   IF #COM_RST              // полный сброс
   THEN
       #LMNR_SIM:=#LMNRSVAL;
       #QLMNUP:=0;
       #QLMNDN:=0;
       #PV:=0.0;
       #ER:=0.0;
       #LMNRS_ON:=0;
       #LMNRSVAL:=0.0;
       #LMNR_SIM:=0.0;
       #sFbPVal:=0.0;
       #sThrOn:=0.0;
       #siImpAus:=0;
       #stImpDauer:=T#0MS;
       #stPausDauer:=T#0MS;
   ELSE
       #Istwert:=INT_TO_REAL(WORD_TO_INT(#PV_PER))*3.616898e-003;
       #Istwert:=#Istwert*#PV_FAC+#PV_OFF;
       IF NOT #PVPER_ON THEN #Istwert:=#PV_IN; END_IF;
       #PV:=#Istwert;
       #ErKp:=#SP_INT-#PV;
       IF    #ErKp < (-#DEADB_W) THEN  #ER:=#ErKp+#DEADB_W;
       ELSIF #ErKp>#DEADB_W      THEN  #ER:=#ErKp-#DEADB_W;
       ELSE  #ER:=0.0; END_IF;
       #ErKp:=#ER*#GAIN;
       #rCycle:=DINT_TO_REAL(TIME_TO_DINT(#CYCLE))/1000.0;
       #rTi:=DINT_TO_REAL(TIME_TO_DINT(#TI))/1000.0;
       IF #rTi<#rCycle*0.5 THEN #rTi:=#rCycle*0.5; END_IF;
       #rMtrTm:=DINT_TO_REAL(TIME_TO_DINT(#MTR_TM))/1000.0;
       #Hvar:=#rTi-ABS(0.01*#ErKp*#rMtrTm);
       IF #Hvar<(#rTi*0.1)THEN #rTi:=#rTi*0.1; ELSE #rTi:=#Hvar; END_IF; 
       IF #LMNS_ON
       THEN
           #sFbPVal:=0.0;
       ELSE 
           IF #siImpAus<>0
           THEN 
               #dInteg:=DINT_TO_REAL(INT_TO_DINT(#siImpAus))*#rCycle/#rMtrTm;
           ELSE
               IF (#ErKp>0.0 AND #LMNR_HS) OR (#ErKp<0.0 AND #LMNR_LS) OR (#TI=T#0MS) 
               THEN
                   #dInteg:=0.0;
               ELSE   
                   #dInteg := (-#ErKp)*#rCycle/#rTi;
               END_IF;
           END_IF;
           #sFbPVal:=#sFbPVal+#dInteg;
           IF #TI=T#0MS
           THEN 
               IF    #sFbPVal>100.0 THEN #sFbPVal:=100.0;
               ELSIF #sFbPVal<0.0   THEN #sFbPVal:=0.0;
               END_IF;
           END_IF;   
       END_IF;       
       #dThrStIn:=#ErKp-#sFbPVal+#DISV;
       #AdapIn1:=#ErKp;
       #AdapIn2:=#sFbPVal;
       #rThrOff:=55.0/#rMtrTm*#rCycle;
       IF #PULSE_TM>#CYCLE
       THEN 
       #Hvar:=DINT_TO_REAL(TIME_TO_DINT(#PULSE_TM))/1000.0;
       ELSE
       #Hvar:=#rCycle;
       END_IF;
       #Hvar:=100.0*#Hvar/#rMtrTm;
       IF NOT(#LMNR_HS OR #LMNR_LS)
       THEN
           IF NOT (#QLMNUP OR #QLMNDN)
           THEN
               IF #TI<>T#0MS
               THEN
                   IF ABS(#AdapIn1)<ABS(#AdapIn2)
                   THEN
                       #sThrOn:=#AdapIn1;
                   ELSE    
                       #sThrOn:=#AdapIn2;
                   END_IF;
               ELSE
                   IF #Istwert=0.0
                   THEN
                       #sThrOn:=#Hvar;
                   ELSE
                       #sThrOn:=ABS(#ErKp)*0.5;
                   END_IF;
               END_IF;
               IF #sThrOn>10.0 THEN #sThrOn:=10.0; END_IF;
               IF #sThrOn<#Hvar THEN #sThrOn:=#Hvar; END_IF;            
           END_IF;           
       ELSE 
           #sThrOn:=#Hvar;
       END_IF;     
       IF (#siImpAus=100 AND #dThrStIn>#rThrOff) OR (#dThrStIn>=#sThrOn)             THEN #iImpEin:=100;
       ELSIF (#siImpAus=-100 AND #dThrStIn<(-#rThrOff)) OR (#dThrStIn<=(-#sThrOn))   THEN #iImpEin:=-100;
       ELSE                                                                          #iImpEin:=0;     
       END_IF;
       IF  #LMNS_ON
       THEN
           IF #LMNUP XOR #LMNDN 
           THEN
               IF #LMNUP
               THEN
                   #iImpEin:=100;
               ELSE
                   #iImpEin:=-100;
               END_IF;
           ELSE
               #iImpEin:=0;
           END_IF;
       END_IF;   
       IF (#iImpEin=100 AND #LMNR_HS) OR (#iImpEin=-100 AND #LMNR_LS) THEN #iImpEin:=0; END_IF;
       IF (#siImpAus=-100 AND #iImpEin=100) OR (#siImpAus=100 AND #iImpEin=-100)THEN #iImpEin:=0; END_IF;
       IF #siImpAus<>#iImpEin
       THEN
           IF #iImpEin=0
           THEN
               IF #stImpDauer<=T#0MS
               THEN
                   #siImpAus:=0;
                   #stPausDauer:=#BREAK_TM;
               END_IF;
           ELSE
               #siImpAus:=#iImpEin;
               #stImpDauer:=#PULSE_TM;
           END_IF;
       END_IF;
       IF #stImpDauer>T#0MS
       THEN
       #stImpDauer:=#stImpDauer-#CYCLE;
       ELSE
       #stImpDauer:=T#0MS;
       END_IF;
       IF #stPausDauer>T#0MS
       THEN
       #stPausDauer:=#stPausDauer-#CYCLE;
       ELSE 
       #stPausDauer:=T#0MS;
       END_IF;
       IF ((#siImpAus=100) AND #LMNR_HS) OR ((#siImpAus=-100) AND #LMNR_LS)
       THEN
         #siImpAus:=0;
         #stImpDauer:=T#0MS;
       END_IF;
       IF NOT #LMNRS_ON
       THEN
           #LmnrSim:=#LMNRSVAL;
       ELSE
           #LmnrSim:=DINT_TO_REAL(INT_TO_DINT(#siImpAus))*#rCycle/#rMtrTm+#LMNR_SIM;
           IF #LmnrSim>=100.0
           THEN
               #LmnrSim:=100.0;
           ELSIF  #LmnrSim<=0.0
           THEN
               #LmnrSim:=0.0;
           END_IF;
       END_IF;
       #LMNR_SIM:=#LmnrSim;
       IF #siImpAus=0
       THEN
              #QLMNUP:=0;
              #QLMNDN:=0;
       ELSIF #siImpAus=100
       THEN
           #QLMNUP:=1;
                 #QLMNDN:=0;
       ELSE
              #QLMNUP:=0;
              #QLMNDN:=1;
       END_IF;
   END_IF;
END_FUNCTION_BLOCK

FUNCTION "03_FC_PID" : Void   // FC3, LAD
{ S7_Optimized_Access := 'FALSE' }
VERSION : 0.1
BEGIN

REGION Network 1
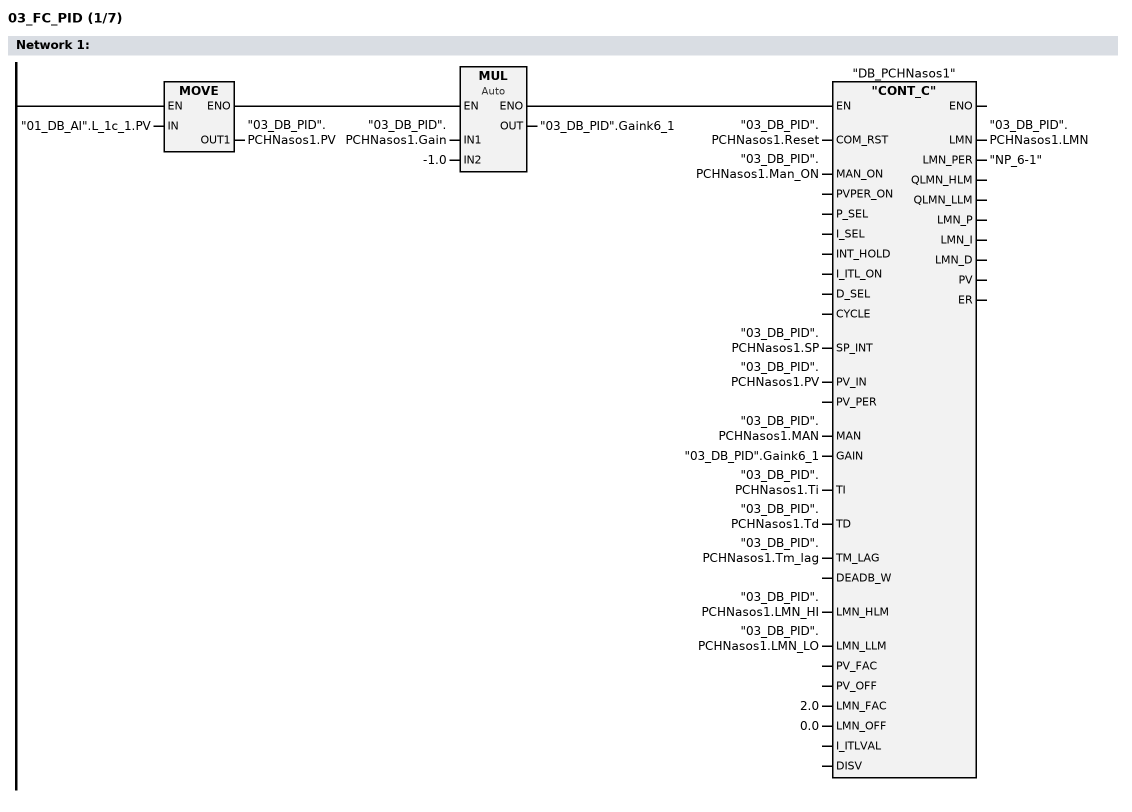
   RUNG wire#powerrail
      Move(in := "01_DB_AI".L_1c_1.PV, out1 => "03_DB_PID".PCHNasos1.PV)
      Mul(in1 := "03_DB_PID".PCHNasos1.Gain, in2 := -1.0, out => "03_DB_PID".Gaink6_1)
      "DB_PCHNasos1"(COM_RST := "03_DB_PID".PCHNasos1.Reset, MAN_ON := "03_DB_PID".PCHNasos1.Man_ON, PVPER_ON :=, P_SEL :=, I_SEL :=, INT_HOLD :=, I_ITL_ON :=, D_SEL :=, CYCLE :=, SP_INT := "03_DB_PID".PCHNasos1.SP, PV_IN := "03_DB_PID".PCHNasos1.PV, PV_PER :=, MAN := "03_DB_PID".PCHNasos1.MAN, GAIN := "03_DB_PID".Gaink6_1, TI := "03_DB_PID".PCHNasos1.Ti, TD := "03_DB_PID".PCHNasos1.Td, TM_LAG := "03_DB_PID".PCHNasos1.Tm_lag, DEADB_W :=, LMN_HLM := "03_DB_PID".PCHNasos1.LMN_HI, LMN_LLM := "03_DB_PID".PCHNasos1.LMN_LO, PV_FAC :=, PV_OFF :=, LMN_FAC := 2.0, LMN_OFF := 0.0, I_ITLVAL :=, DISV :=, LMN => "03_DB_PID".PCHNasos1.LMN, LMN_PER => "NP_6-1", QLMN_HLM =>, QLMN_LLM =>, LMN_P =>, LMN_I =>, LMN_D =>, PV =>, ER =>)
   END_RUNG
   // the same network as SCL:
   "03_DB_PID".PCHNasos1.PV := "01_DB_AI".L_1c_1.PV;
   "03_DB_PID".Gaink6_1 := "03_DB_PID".PCHNasos1.Gain * (-1.0);
   "DB_PCHNasos1"(COM_RST := "03_DB_PID".PCHNasos1.Reset,   // "CONT_C"
                  MAN_ON := "03_DB_PID".PCHNasos1.Man_ON,
                  SP_INT := "03_DB_PID".PCHNasos1.SP,
                  PV_IN := "03_DB_PID".PCHNasos1.PV,
                  MAN := "03_DB_PID".PCHNasos1.MAN,
                  GAIN := "03_DB_PID".Gaink6_1,
                  TI := "03_DB_PID".PCHNasos1.Ti,
                  TD := "03_DB_PID".PCHNasos1.Td,
                  TM_LAG := "03_DB_PID".PCHNasos1.Tm_lag,
                  LMN_HLM := "03_DB_PID".PCHNasos1.LMN_HI,
                  LMN_LLM := "03_DB_PID".PCHNasos1.LMN_LO,
                  LMN_FAC := 2.0,
                  LMN_OFF := 0.0,
                  LMN => "03_DB_PID".PCHNasos1.LMN,
                  LMN_PER => "NP_6-1");
END_REGION

REGION Network 2
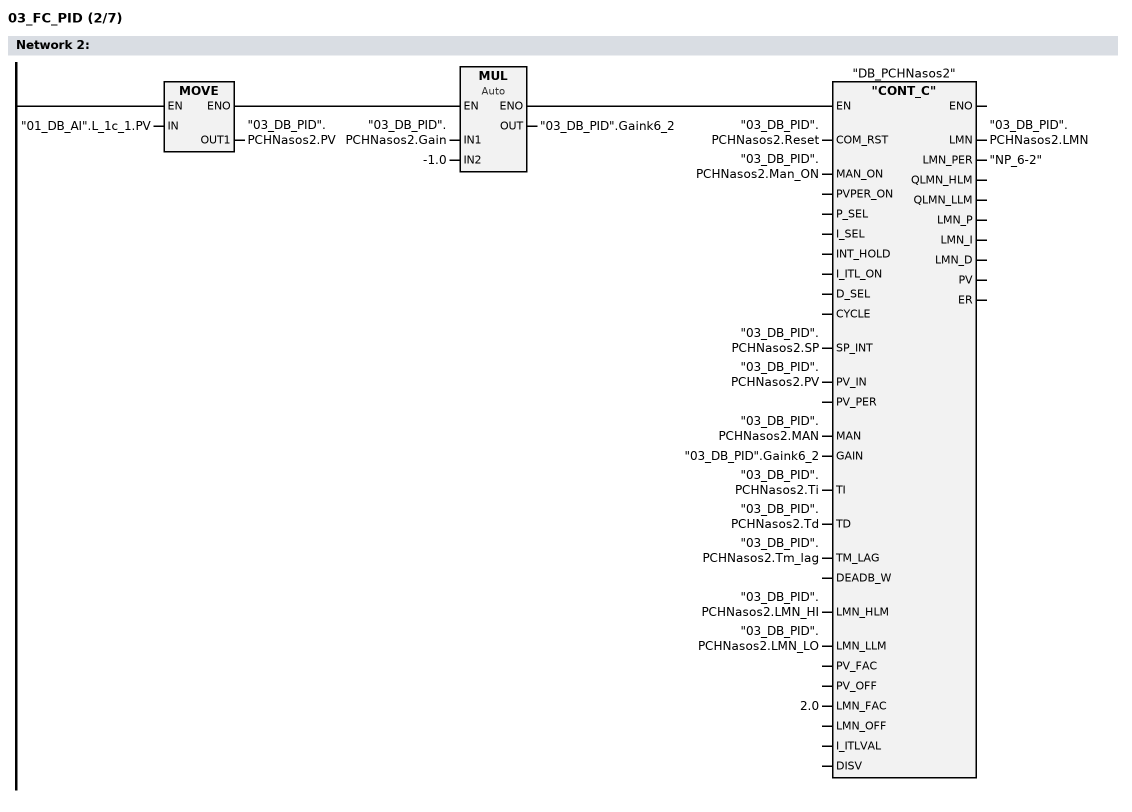
   RUNG wire#powerrail
      Move(in := "01_DB_AI".L_1c_1.PV, out1 => "03_DB_PID".PCHNasos2.PV)
      Mul(in1 := "03_DB_PID".PCHNasos2.Gain, in2 := -1.0, out => "03_DB_PID".Gaink6_2)
      "DB_PCHNasos2"(COM_RST := "03_DB_PID".PCHNasos2.Reset, MAN_ON := "03_DB_PID".PCHNasos2.Man_ON, PVPER_ON :=, P_SEL :=, I_SEL :=, INT_HOLD :=, I_ITL_ON :=, D_SEL :=, CYCLE :=, SP_INT := "03_DB_PID".PCHNasos2.SP, PV_IN := "03_DB_PID".PCHNasos2.PV, PV_PER :=, MAN := "03_DB_PID".PCHNasos2.MAN, GAIN := "03_DB_PID".Gaink6_2, TI := "03_DB_PID".PCHNasos2.Ti, TD := "03_DB_PID".PCHNasos2.Td, TM_LAG := "03_DB_PID".PCHNasos2.Tm_lag, DEADB_W :=, LMN_HLM := "03_DB_PID".PCHNasos2.LMN_HI, LMN_LLM := "03_DB_PID".PCHNasos2.LMN_LO, PV_FAC :=, PV_OFF :=, LMN_FAC := 2.0, LMN_OFF :=, I_ITLVAL :=, DISV :=, LMN => "03_DB_PID".PCHNasos2.LMN, LMN_PER => "NP_6-2", QLMN_HLM =>, QLMN_LLM =>, LMN_P =>, LMN_I =>, LMN_D =>, PV =>, ER =>)
   END_RUNG
   // the same network as SCL:
   "03_DB_PID".PCHNasos2.PV := "01_DB_AI".L_1c_1.PV;
   "03_DB_PID".Gaink6_2 := "03_DB_PID".PCHNasos2.Gain * (-1.0);
   "DB_PCHNasos2"(COM_RST := "03_DB_PID".PCHNasos2.Reset,   // "CONT_C"
                  MAN_ON := "03_DB_PID".PCHNasos2.Man_ON,
                  SP_INT := "03_DB_PID".PCHNasos2.SP,
                  PV_IN := "03_DB_PID".PCHNasos2.PV,
                  MAN := "03_DB_PID".PCHNasos2.MAN,
                  GAIN := "03_DB_PID".Gaink6_2,
                  TI := "03_DB_PID".PCHNasos2.Ti,
                  TD := "03_DB_PID".PCHNasos2.Td,
                  TM_LAG := "03_DB_PID".PCHNasos2.Tm_lag,
                  LMN_HLM := "03_DB_PID".PCHNasos2.LMN_HI,
                  LMN_LLM := "03_DB_PID".PCHNasos2.LMN_LO,
                  LMN_FAC := 2.0,
                  LMN => "03_DB_PID".PCHNasos2.LMN,
                  LMN_PER => "NP_6-2");
END_REGION

REGION Network 3
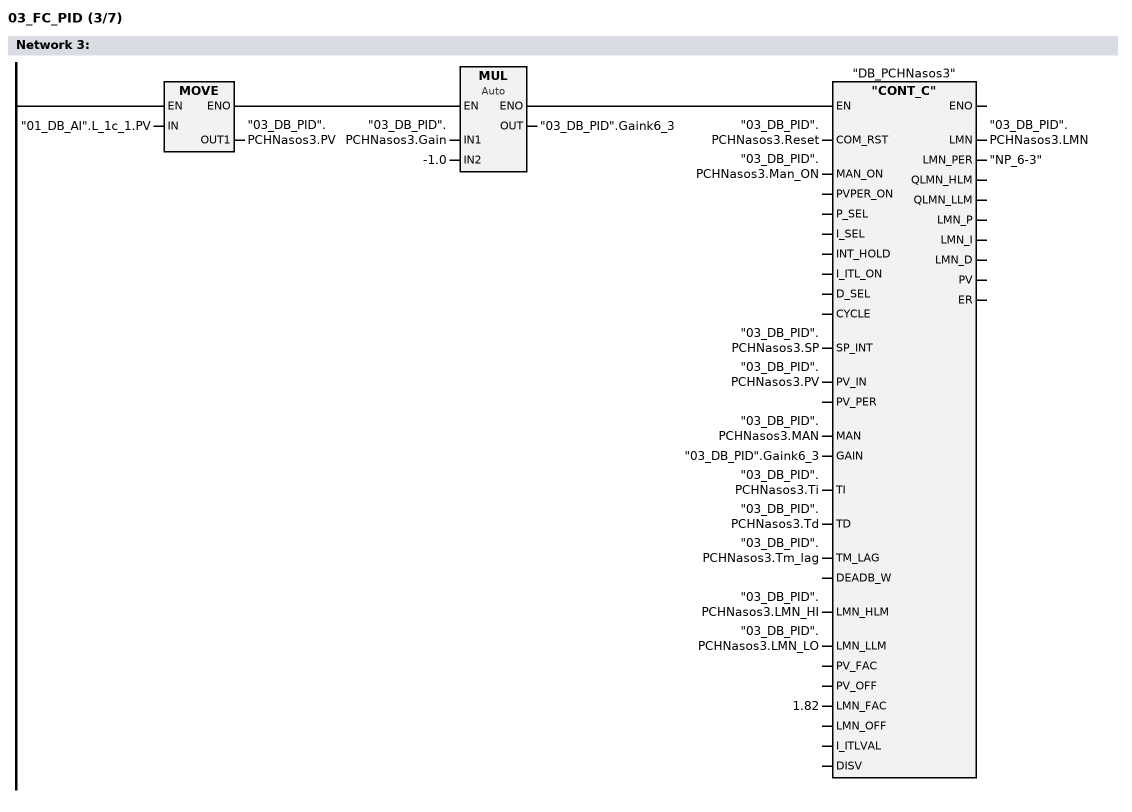
   RUNG wire#powerrail
      Move(in := "01_DB_AI".L_1c_1.PV, out1 => "03_DB_PID".PCHNasos3.PV)
      Mul(in1 := "03_DB_PID".PCHNasos3.Gain, in2 := -1.0, out => "03_DB_PID".Gaink6_3)
      "DB_PCHNasos3"(COM_RST := "03_DB_PID".PCHNasos3.Reset, MAN_ON := "03_DB_PID".PCHNasos3.Man_ON, PVPER_ON :=, P_SEL :=, I_SEL :=, INT_HOLD :=, I_ITL_ON :=, D_SEL :=, CYCLE :=, SP_INT := "03_DB_PID".PCHNasos3.SP, PV_IN := "03_DB_PID".PCHNasos3.PV, PV_PER :=, MAN := "03_DB_PID".PCHNasos3.MAN, GAIN := "03_DB_PID".Gaink6_3, TI := "03_DB_PID".PCHNasos3.Ti, TD := "03_DB_PID".PCHNasos3.Td, TM_LAG := "03_DB_PID".PCHNasos3.Tm_lag, DEADB_W :=, LMN_HLM := "03_DB_PID".PCHNasos3.LMN_HI, LMN_LLM := "03_DB_PID".PCHNasos3.LMN_LO, PV_FAC :=, PV_OFF :=, LMN_FAC := 1.82, LMN_OFF :=, I_ITLVAL :=, DISV :=, LMN => "03_DB_PID".PCHNasos3.LMN, LMN_PER => "NP_6-3", QLMN_HLM =>, QLMN_LLM =>, LMN_P =>, LMN_I =>, LMN_D =>, PV =>, ER =>)
   END_RUNG
   // the same network as SCL:
   "03_DB_PID".PCHNasos3.PV := "01_DB_AI".L_1c_1.PV;
   "03_DB_PID".Gaink6_3 := "03_DB_PID".PCHNasos3.Gain * (-1.0);
   "DB_PCHNasos3"(COM_RST := "03_DB_PID".PCHNasos3.Reset,   // "CONT_C"
                  MAN_ON := "03_DB_PID".PCHNasos3.Man_ON,
                  SP_INT := "03_DB_PID".PCHNasos3.SP,
                  PV_IN := "03_DB_PID".PCHNasos3.PV,
                  MAN := "03_DB_PID".PCHNasos3.MAN,
                  GAIN := "03_DB_PID".Gaink6_3,
                  TI := "03_DB_PID".PCHNasos3.Ti,
                  TD := "03_DB_PID".PCHNasos3.Td,
                  TM_LAG := "03_DB_PID".PCHNasos3.Tm_lag,
                  LMN_HLM := "03_DB_PID".PCHNasos3.LMN_HI,
                  LMN_LLM := "03_DB_PID".PCHNasos3.LMN_LO,
                  LMN_FAC := 1.82,
                  LMN => "03_DB_PID".PCHNasos3.LMN,
                  LMN_PER => "NP_6-3");
END_REGION

REGION Network 4
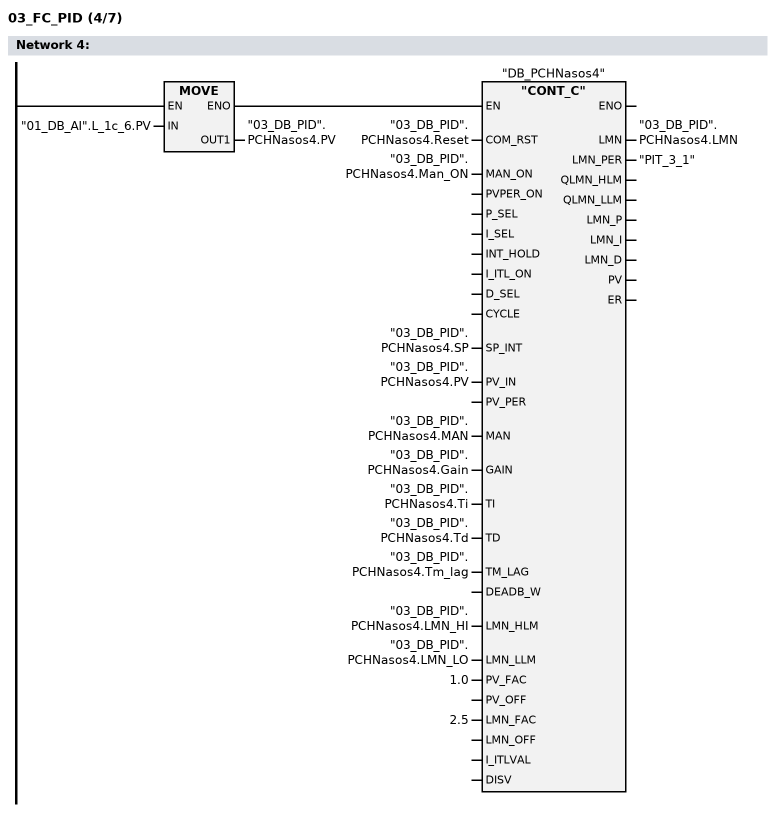
   RUNG wire#powerrail
      Move(in := "01_DB_AI".L_1c_6.PV, out1 => "03_DB_PID".PCHNasos4.PV)
      "DB_PCHNasos4"(COM_RST := "03_DB_PID".PCHNasos4.Reset, MAN_ON := "03_DB_PID".PCHNasos4.Man_ON, PVPER_ON :=, P_SEL :=, I_SEL :=, INT_HOLD :=, I_ITL_ON :=, D_SEL :=, CYCLE :=, SP_INT := "03_DB_PID".PCHNasos4.SP, PV_IN := "03_DB_PID".PCHNasos4.PV, PV_PER :=, MAN := "03_DB_PID".PCHNasos4.MAN, GAIN := "03_DB_PID".PCHNasos4.Gain, TI := "03_DB_PID".PCHNasos4.Ti, TD := "03_DB_PID".PCHNasos4.Td, TM_LAG := "03_DB_PID".PCHNasos4.Tm_lag, DEADB_W :=, LMN_HLM := "03_DB_PID".PCHNasos4.LMN_HI, LMN_LLM := "03_DB_PID".PCHNasos4.LMN_LO, PV_FAC := 1.0, PV_OFF :=, LMN_FAC := 2.5, LMN_OFF :=, I_ITLVAL :=, DISV :=, LMN => "03_DB_PID".PCHNasos4.LMN, LMN_PER => "PIT_3_1", QLMN_HLM =>, QLMN_LLM =>, LMN_P =>, LMN_I =>, LMN_D =>, PV =>, ER =>)
   END_RUNG
   // the same network as SCL:
   "03_DB_PID".PCHNasos4.PV := "01_DB_AI".L_1c_6.PV;
   "DB_PCHNasos4"(COM_RST := "03_DB_PID".PCHNasos4.Reset,   // "CONT_C"
                  MAN_ON := "03_DB_PID".PCHNasos4.Man_ON,
                  SP_INT := "03_DB_PID".PCHNasos4.SP,
                  PV_IN := "03_DB_PID".PCHNasos4.PV,
                  MAN := "03_DB_PID".PCHNasos4.MAN,
                  GAIN := "03_DB_PID".PCHNasos4.Gain,
                  TI := "03_DB_PID".PCHNasos4.Ti,
                  TD := "03_DB_PID".PCHNasos4.Td,
                  TM_LAG := "03_DB_PID".PCHNasos4.Tm_lag,
                  LMN_HLM := "03_DB_PID".PCHNasos4.LMN_HI,
                  LMN_LLM := "03_DB_PID".PCHNasos4.LMN_LO,
                  PV_FAC := 1.0,
                  LMN_FAC := 2.5,
                  LMN => "03_DB_PID".PCHNasos4.LMN,
                  LMN_PER => "PIT_3_1");
END_REGION

REGION Network 5
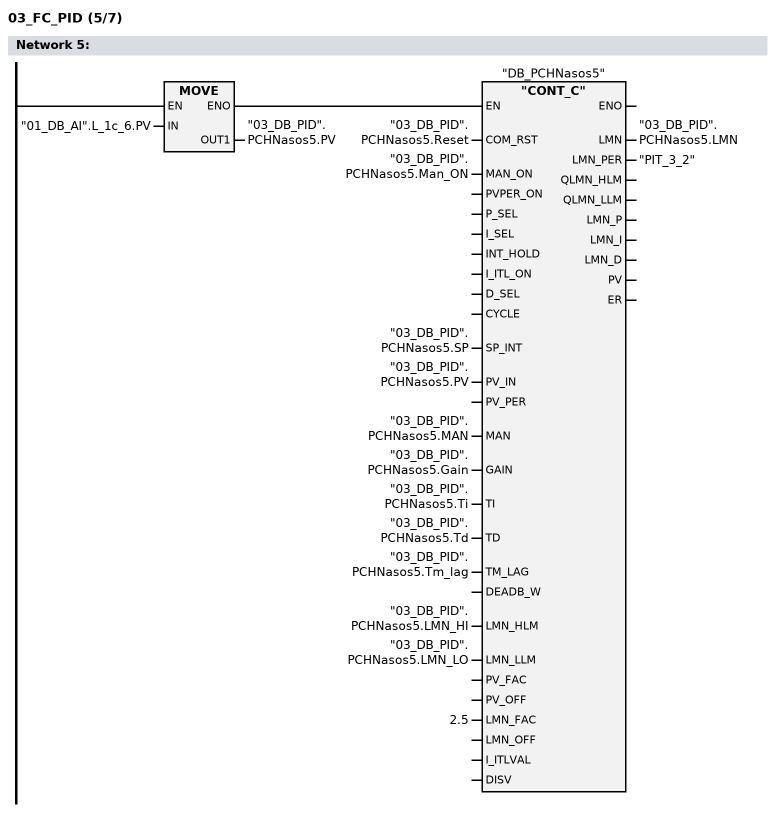
   RUNG wire#powerrail
      Move(in := "01_DB_AI".L_1c_6.PV, out1 => "03_DB_PID".PCHNasos5.PV)
      "DB_PCHNasos5"(COM_RST := "03_DB_PID".PCHNasos5.Reset, MAN_ON := "03_DB_PID".PCHNasos5.Man_ON, PVPER_ON :=, P_SEL :=, I_SEL :=, INT_HOLD :=, I_ITL_ON :=, D_SEL :=, CYCLE :=, SP_INT := "03_DB_PID".PCHNasos5.SP, PV_IN := "03_DB_PID".PCHNasos5.PV, PV_PER :=, MAN := "03_DB_PID".PCHNasos5.MAN, GAIN := "03_DB_PID".PCHNasos5.Gain, TI := "03_DB_PID".PCHNasos5.Ti, TD := "03_DB_PID".PCHNasos5.Td, TM_LAG := "03_DB_PID".PCHNasos5.Tm_lag, DEADB_W :=, LMN_HLM := "03_DB_PID".PCHNasos5.LMN_HI, LMN_LLM := "03_DB_PID".PCHNasos5.LMN_LO, PV_FAC :=, PV_OFF :=, LMN_FAC := 2.5, LMN_OFF :=, I_ITLVAL :=, DISV :=, LMN => "03_DB_PID".PCHNasos5.LMN, LMN_PER => "PIT_3_2", QLMN_HLM =>, QLMN_LLM =>, LMN_P =>, LMN_I =>, LMN_D =>, PV =>, ER =>)
   END_RUNG
   // the same network as SCL:
   "03_DB_PID".PCHNasos5.PV := "01_DB_AI".L_1c_6.PV;
   "DB_PCHNasos5"(COM_RST := "03_DB_PID".PCHNasos5.Reset,   // "CONT_C"
                  MAN_ON := "03_DB_PID".PCHNasos5.Man_ON,
                  SP_INT := "03_DB_PID".PCHNasos5.SP,
                  PV_IN := "03_DB_PID".PCHNasos5.PV,
                  MAN := "03_DB_PID".PCHNasos5.MAN,
                  GAIN := "03_DB_PID".PCHNasos5.Gain,
                  TI := "03_DB_PID".PCHNasos5.Ti,
                  TD := "03_DB_PID".PCHNasos5.Td,
                  TM_LAG := "03_DB_PID".PCHNasos5.Tm_lag,
                  LMN_HLM := "03_DB_PID".PCHNasos5.LMN_HI,
                  LMN_LLM := "03_DB_PID".PCHNasos5.LMN_LO,
                  LMN_FAC := 2.5,
                  LMN => "03_DB_PID".PCHNasos5.LMN,
                  LMN_PER => "PIT_3_2");
END_REGION

REGION Network 6
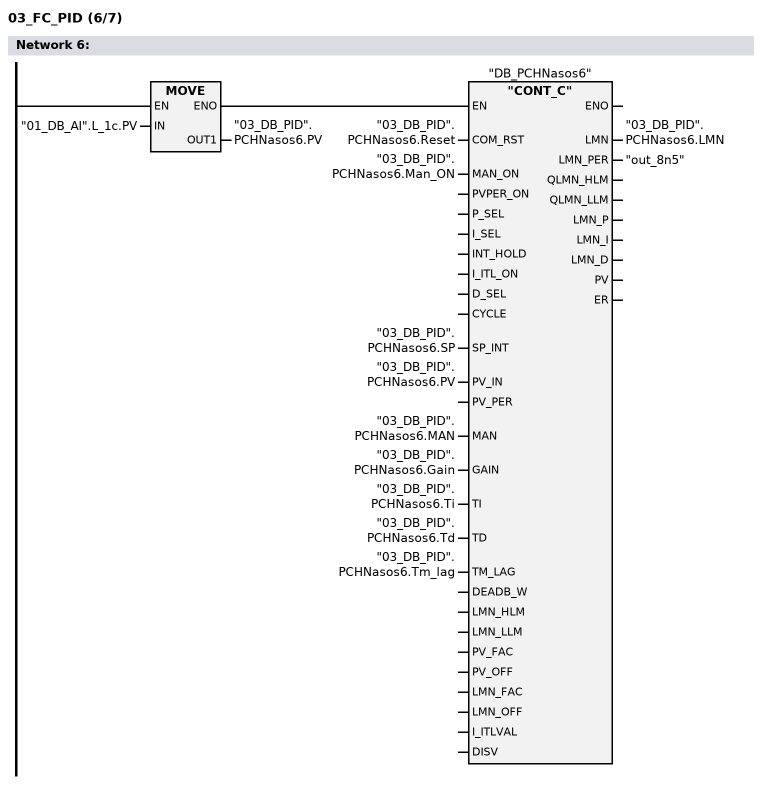
   RUNG wire#powerrail
      Move(in := "01_DB_AI".L_1c.PV, out1 => "03_DB_PID".PCHNasos6.PV)
      "DB_PCHNasos6"(COM_RST := "03_DB_PID".PCHNasos6.Reset, MAN_ON := "03_DB_PID".PCHNasos6.Man_ON, PVPER_ON :=, P_SEL :=, I_SEL :=, INT_HOLD :=, I_ITL_ON :=, D_SEL :=, CYCLE :=, SP_INT := "03_DB_PID".PCHNasos6.SP, PV_IN := "03_DB_PID".PCHNasos6.PV, PV_PER :=, MAN := "03_DB_PID".PCHNasos6.MAN, GAIN := "03_DB_PID".PCHNasos6.Gain, TI := "03_DB_PID".PCHNasos6.Ti, TD := "03_DB_PID".PCHNasos6.Td, TM_LAG := "03_DB_PID".PCHNasos6.Tm_lag, DEADB_W :=, LMN_HLM :=, LMN_LLM :=, PV_FAC :=, PV_OFF :=, LMN_FAC :=, LMN_OFF :=, I_ITLVAL :=, DISV :=, LMN => "03_DB_PID".PCHNasos6.LMN, LMN_PER => "out_8n5", QLMN_HLM =>, QLMN_LLM =>, LMN_P =>, LMN_I =>, LMN_D =>, PV =>, ER =>)
   END_RUNG
   // the same network as SCL:
   "03_DB_PID".PCHNasos6.PV := "01_DB_AI".L_1c.PV;
   "DB_PCHNasos6"(COM_RST := "03_DB_PID".PCHNasos6.Reset,   // "CONT_C"
                  MAN_ON := "03_DB_PID".PCHNasos6.Man_ON,
                  SP_INT := "03_DB_PID".PCHNasos6.SP,
                  PV_IN := "03_DB_PID".PCHNasos6.PV,
                  MAN := "03_DB_PID".PCHNasos6.MAN,
                  GAIN := "03_DB_PID".PCHNasos6.Gain,
                  TI := "03_DB_PID".PCHNasos6.Ti,
                  TD := "03_DB_PID".PCHNasos6.Td,
                  TM_LAG := "03_DB_PID".PCHNasos6.Tm_lag,
                  LMN => "03_DB_PID".PCHNasos6.LMN,
                  LMN_PER => "out_8n5");
END_REGION

REGION Network 7
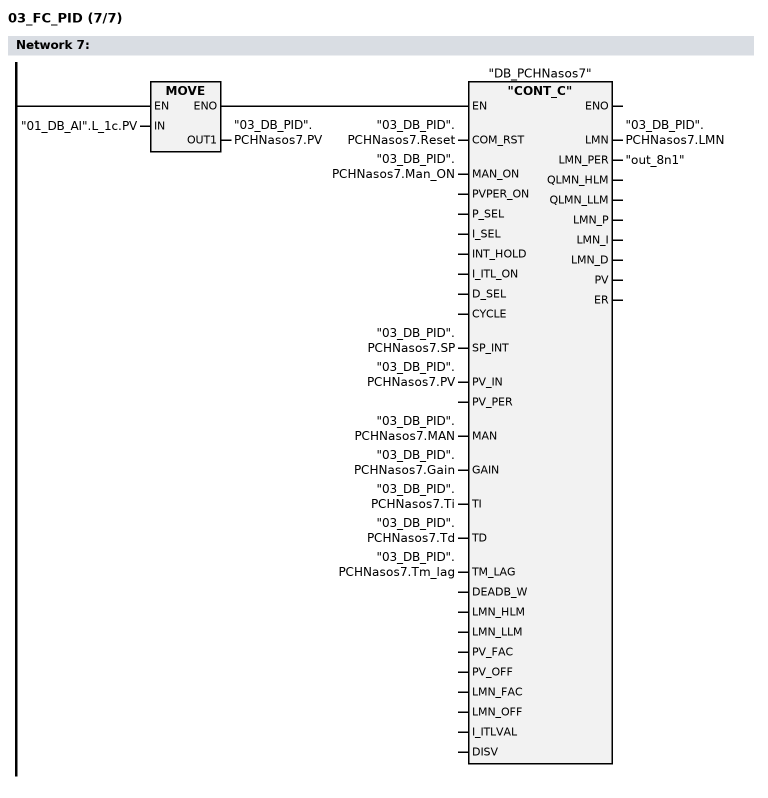
   RUNG wire#powerrail
      Move(in := "01_DB_AI".L_1c.PV, out1 => "03_DB_PID".PCHNasos7.PV)
      "DB_PCHNasos7"(COM_RST := "03_DB_PID".PCHNasos7.Reset, MAN_ON := "03_DB_PID".PCHNasos7.Man_ON, PVPER_ON :=, P_SEL :=, I_SEL :=, INT_HOLD :=, I_ITL_ON :=, D_SEL :=, CYCLE :=, SP_INT := "03_DB_PID".PCHNasos7.SP, PV_IN := "03_DB_PID".PCHNasos7.PV, PV_PER :=, MAN := "03_DB_PID".PCHNasos7.MAN, GAIN := "03_DB_PID".PCHNasos7.Gain, TI := "03_DB_PID".PCHNasos7.Ti, TD := "03_DB_PID".PCHNasos7.Td, TM_LAG := "03_DB_PID".PCHNasos7.Tm_lag, DEADB_W :=, LMN_HLM :=, LMN_LLM :=, PV_FAC :=, PV_OFF :=, LMN_FAC :=, LMN_OFF :=, I_ITLVAL :=, DISV :=, LMN => "03_DB_PID".PCHNasos7.LMN, LMN_PER => "out_8n1", QLMN_HLM =>, QLMN_LLM =>, LMN_P =>, LMN_I =>, LMN_D =>, PV =>, ER =>)
   END_RUNG
   // the same network as SCL:
   "03_DB_PID".PCHNasos7.PV := "01_DB_AI".L_1c.PV;
   "DB_PCHNasos7"(COM_RST := "03_DB_PID".PCHNasos7.Reset,   // "CONT_C"
                  MAN_ON := "03_DB_PID".PCHNasos7.Man_ON,
                  SP_INT := "03_DB_PID".PCHNasos7.SP,
                  PV_IN := "03_DB_PID".PCHNasos7.PV,
                  MAN := "03_DB_PID".PCHNasos7.MAN,
                  GAIN := "03_DB_PID".PCHNasos7.Gain,
                  TI := "03_DB_PID".PCHNasos7.Ti,
                  TD := "03_DB_PID".PCHNasos7.Td,
                  TM_LAG := "03_DB_PID".PCHNasos7.Tm_lag,
                  LMN => "03_DB_PID".PCHNasos7.LMN,
                  LMN_PER => "out_8n1");
END_REGION
END_FUNCTION

FUNCTION "06_FC_MOTORS" : Void   // FC6, LAD
{ S7_Optimized_Access := 'TRUE' }
VERSION : 0.1
   VAR_TEMP
      LocRem : Bool;
      out : Bool;
   END_VAR
   VAR_TEMP   // added for the SCL form of the ladder/FBD networks
      _w1 : Bool;
   END_VAR
BEGIN

REGION Network 1
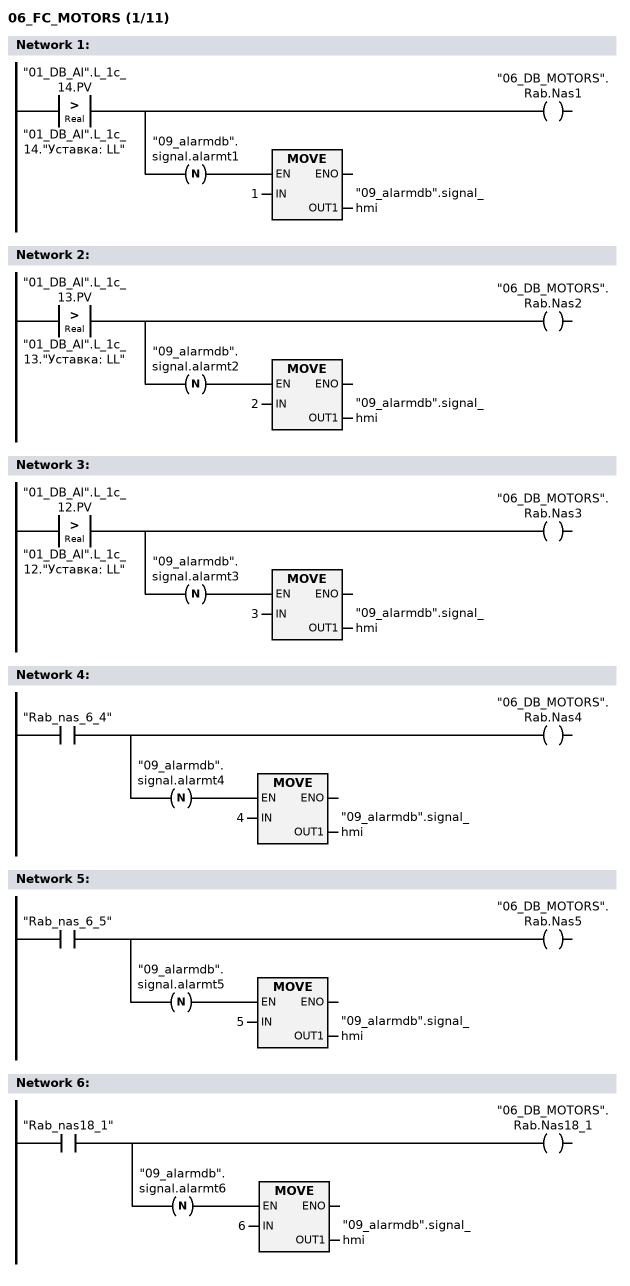
   RUNG wire#powerrail
      { S7_Templates := "SrcType := Real" } GT_Contact(in1 := "01_DB_AI".L_1c_14.PV, in2 := "01_DB_AI".L_1c_14."Уставка: LL")
      wire#w1
      Coil( "06_DB_MOTORS".Rab.Nas1 )
   END_RUNG
   RUNG wire#w1
      N_Trig( "09_alarmdb".signal.alarmt1 )
      Move(in := 1, out1 => "09_alarmdb".signal_hmi)
   END_RUNG
   // the same network as SCL:
   "06_DB_MOTORS".Rab.Nas1 := "01_DB_AI".L_1c_14.PV > "01_DB_AI".L_1c_14."Уставка: LL";
   #_w1 := NOT "06_DB_MOTORS".Rab.Nas1 AND "09_alarmdb".signal.alarmt1;   // falling edge
   "09_alarmdb".signal.alarmt1 := "06_DB_MOTORS".Rab.Nas1;
   IF #_w1 THEN "09_alarmdb".signal_hmi := 1; END_IF;
END_REGION

REGION Network 2
   RUNG wire#powerrail
      { S7_Templates := "SrcType := Real" } GT_Contact(in1 := "01_DB_AI".L_1c_13.PV, in2 := "01_DB_AI".L_1c_13."Уставка: LL")
      wire#w1
      Coil( "06_DB_MOTORS".Rab.Nas2 )
   END_RUNG
   RUNG wire#w1
      N_Trig( "09_alarmdb".signal.alarmt2 )
      Move(in := 2, out1 => "09_alarmdb".signal_hmi)
   END_RUNG
   // the same network as SCL:
   "06_DB_MOTORS".Rab.Nas2 := "01_DB_AI".L_1c_13.PV > "01_DB_AI".L_1c_13."Уставка: LL";
   #_w1 := NOT "06_DB_MOTORS".Rab.Nas2 AND "09_alarmdb".signal.alarmt2;   // falling edge
   "09_alarmdb".signal.alarmt2 := "06_DB_MOTORS".Rab.Nas2;
   IF #_w1 THEN "09_alarmdb".signal_hmi := 2; END_IF;
END_REGION

REGION Network 3
   RUNG wire#powerrail
      { S7_Templates := "SrcType := Real" } GT_Contact(in1 := "01_DB_AI".L_1c_12.PV, in2 := "01_DB_AI".L_1c_12."Уставка: LL")
      wire#w1
      Coil( "06_DB_MOTORS".Rab.Nas3 )
   END_RUNG
   RUNG wire#w1
      N_Trig( "09_alarmdb".signal.alarmt3 )
      Move(in := 3, out1 => "09_alarmdb".signal_hmi)
   END_RUNG
   // the same network as SCL:
   "06_DB_MOTORS".Rab.Nas3 := "01_DB_AI".L_1c_12.PV > "01_DB_AI".L_1c_12."Уставка: LL";
   #_w1 := NOT "06_DB_MOTORS".Rab.Nas3 AND "09_alarmdb".signal.alarmt3;   // falling edge
   "09_alarmdb".signal.alarmt3 := "06_DB_MOTORS".Rab.Nas3;
   IF #_w1 THEN "09_alarmdb".signal_hmi := 3; END_IF;
END_REGION

REGION Network 4
   RUNG wire#powerrail
      Contact( "Rab_nas_6_4" )
      wire#w1
      Coil( "06_DB_MOTORS".Rab.Nas4 )
   END_RUNG
   RUNG wire#w1
      N_Trig( "09_alarmdb".signal.alarmt4 )
      Move(in := 4, out1 => "09_alarmdb".signal_hmi)
   END_RUNG
   // the same network as SCL:
   "06_DB_MOTORS".Rab.Nas4 := "Rab_nas_6_4";
   #_w1 := NOT "Rab_nas_6_4" AND "09_alarmdb".signal.alarmt4;   // falling edge
   "09_alarmdb".signal.alarmt4 := "Rab_nas_6_4";
   IF #_w1 THEN "09_alarmdb".signal_hmi := 4; END_IF;
END_REGION

REGION Network 5
   RUNG wire#powerrail
      Contact( "Rab_nas_6_5" )
      wire#w1
      Coil( "06_DB_MOTORS".Rab.Nas5 )
   END_RUNG
   RUNG wire#w1
      N_Trig( "09_alarmdb".signal.alarmt5 )
      Move(in := 5, out1 => "09_alarmdb".signal_hmi)
   END_RUNG
   // the same network as SCL:
   "06_DB_MOTORS".Rab.Nas5 := "Rab_nas_6_5";
   #_w1 := NOT "Rab_nas_6_5" AND "09_alarmdb".signal.alarmt5;   // falling edge
   "09_alarmdb".signal.alarmt5 := "Rab_nas_6_5";
   IF #_w1 THEN "09_alarmdb".signal_hmi := 5; END_IF;
END_REGION

REGION Network 6
   RUNG wire#powerrail
      Contact( "Rab_nas18_1" )
      wire#w1
      Coil( "06_DB_MOTORS".Rab.Nas18_1 )
   END_RUNG
   RUNG wire#w1
      N_Trig( "09_alarmdb".signal.alarmt6 )
      Move(in := 6, out1 => "09_alarmdb".signal_hmi)
   END_RUNG
   // the same network as SCL:
   "06_DB_MOTORS".Rab.Nas18_1 := "Rab_nas18_1";
   #_w1 := NOT "Rab_nas18_1" AND "09_alarmdb".signal.alarmt6;   // falling edge
   "09_alarmdb".signal.alarmt6 := "Rab_nas18_1";
   IF #_w1 THEN "09_alarmdb".signal_hmi := 6; END_IF;
END_REGION

REGION Network 7
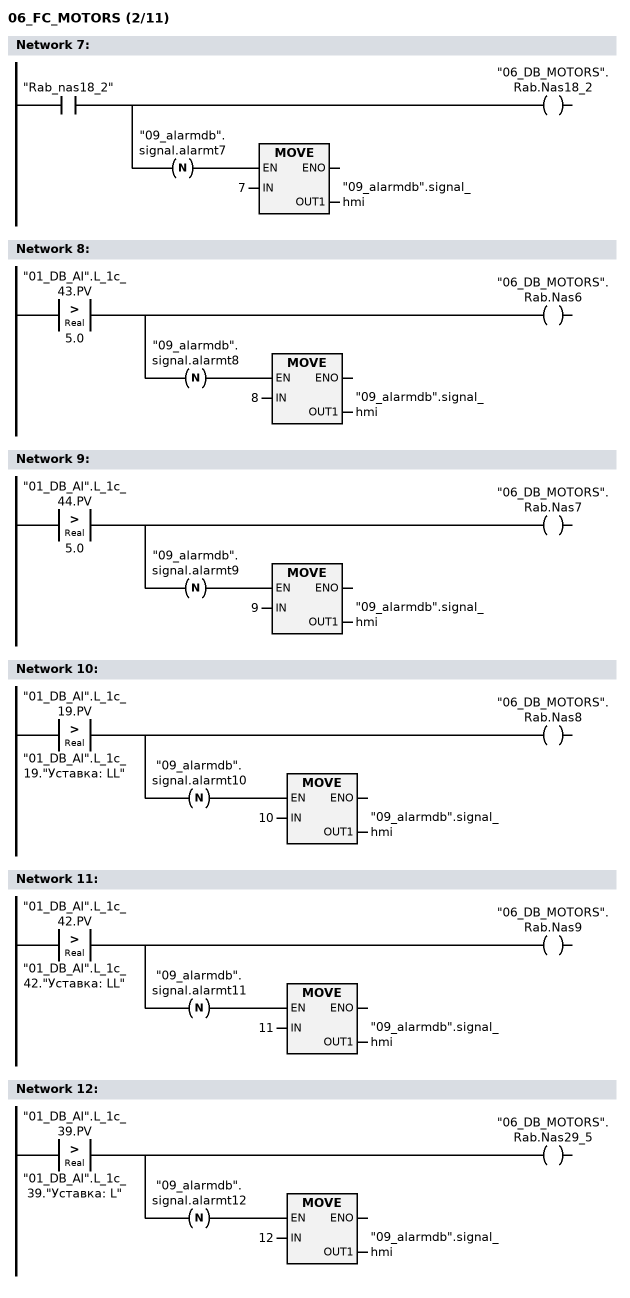
   RUNG wire#powerrail
      Contact( "Rab_nas18_2" )
      wire#w1
      Coil( "06_DB_MOTORS".Rab.Nas18_2 )
   END_RUNG
   RUNG wire#w1
      N_Trig( "09_alarmdb".signal.alarmt7 )
      Move(in := 7, out1 => "09_alarmdb".signal_hmi)
   END_RUNG
   // the same network as SCL:
   "06_DB_MOTORS".Rab.Nas18_2 := "Rab_nas18_2";
   #_w1 := NOT "Rab_nas18_2" AND "09_alarmdb".signal.alarmt7;   // falling edge
   "09_alarmdb".signal.alarmt7 := "Rab_nas18_2";
   IF #_w1 THEN "09_alarmdb".signal_hmi := 7; END_IF;
END_REGION

REGION Network 8
   RUNG wire#powerrail
      { S7_Templates := "SrcType := Real" } GT_Contact(in1 := "01_DB_AI".L_1c_43.PV, in2 := 5.0)
      wire#w1
      Coil( "06_DB_MOTORS".Rab.Nas6 )
   END_RUNG
   RUNG wire#w1
      N_Trig( "09_alarmdb".signal.alarmt8 )
      Move(in := 8, out1 => "09_alarmdb".signal_hmi)
   END_RUNG
   // the same network as SCL:
   "06_DB_MOTORS".Rab.Nas6 := "01_DB_AI".L_1c_43.PV > 5.0;
   #_w1 := NOT "06_DB_MOTORS".Rab.Nas6 AND "09_alarmdb".signal.alarmt8;   // falling edge
   "09_alarmdb".signal.alarmt8 := "06_DB_MOTORS".Rab.Nas6;
   IF #_w1 THEN "09_alarmdb".signal_hmi := 8; END_IF;
END_REGION

REGION Network 9
   RUNG wire#powerrail
      { S7_Templates := "SrcType := Real" } GT_Contact(in1 := "01_DB_AI".L_1c_44.PV, in2 := 5.0)
      wire#w1
      Coil( "06_DB_MOTORS".Rab.Nas7 )
   END_RUNG
   RUNG wire#w1
      N_Trig( "09_alarmdb".signal.alarmt9 )
      Move(in := 9, out1 => "09_alarmdb".signal_hmi)
   END_RUNG
   // the same network as SCL:
   "06_DB_MOTORS".Rab.Nas7 := "01_DB_AI".L_1c_44.PV > 5.0;
   #_w1 := NOT "06_DB_MOTORS".Rab.Nas7 AND "09_alarmdb".signal.alarmt9;   // falling edge
   "09_alarmdb".signal.alarmt9 := "06_DB_MOTORS".Rab.Nas7;
   IF #_w1 THEN "09_alarmdb".signal_hmi := 9; END_IF;
END_REGION

REGION Network 10
   RUNG wire#powerrail
      { S7_Templates := "SrcType := Real" } GT_Contact(in1 := "01_DB_AI".L_1c_19.PV, in2 := "01_DB_AI".L_1c_19."Уставка: LL")
      wire#w1
      Coil( "06_DB_MOTORS".Rab.Nas8 )
   END_RUNG
   RUNG wire#w1
      N_Trig( "09_alarmdb".signal.alarmt10 )
      Move(in := 10, out1 => "09_alarmdb".signal_hmi)
   END_RUNG
   // the same network as SCL:
   "06_DB_MOTORS".Rab.Nas8 := "01_DB_AI".L_1c_19.PV > "01_DB_AI".L_1c_19."Уставка: LL";
   #_w1 := NOT "06_DB_MOTORS".Rab.Nas8 AND "09_alarmdb".signal.alarmt10;   // falling edge
   "09_alarmdb".signal.alarmt10 := "06_DB_MOTORS".Rab.Nas8;
   IF #_w1 THEN "09_alarmdb".signal_hmi := 10; END_IF;
END_REGION

REGION Network 11
   RUNG wire#powerrail
      { S7_Templates := "SrcType := Real" } GT_Contact(in1 := "01_DB_AI".L_1c_42.PV, in2 := "01_DB_AI".L_1c_42."Уставка: LL")
      wire#w1
      Coil( "06_DB_MOTORS".Rab.Nas9 )
   END_RUNG
   RUNG wire#w1
      N_Trig( "09_alarmdb".signal.alarmt11 )
      Move(in := 11, out1 => "09_alarmdb".signal_hmi)
   END_RUNG
   // the same network as SCL:
   "06_DB_MOTORS".Rab.Nas9 := "01_DB_AI".L_1c_42.PV > "01_DB_AI".L_1c_42."Уставка: LL";
   #_w1 := NOT "06_DB_MOTORS".Rab.Nas9 AND "09_alarmdb".signal.alarmt11;   // falling edge
   "09_alarmdb".signal.alarmt11 := "06_DB_MOTORS".Rab.Nas9;
   IF #_w1 THEN "09_alarmdb".signal_hmi := 11; END_IF;
END_REGION

REGION Network 12
   RUNG wire#powerrail
      { S7_Templates := "SrcType := Real" } GT_Contact(in1 := "01_DB_AI".L_1c_39.PV, in2 := "01_DB_AI".L_1c_39."Уставка: L")
      wire#w1
      Coil( "06_DB_MOTORS".Rab.Nas29_5 )
   END_RUNG
   RUNG wire#w1
      N_Trig( "09_alarmdb".signal.alarmt12 )
      Move(in := 12, out1 => "09_alarmdb".signal_hmi)
   END_RUNG
   // the same network as SCL:
   "06_DB_MOTORS".Rab.Nas29_5 := "01_DB_AI".L_1c_39.PV > "01_DB_AI".L_1c_39."Уставка: L";
   #_w1 := NOT "06_DB_MOTORS".Rab.Nas29_5 AND "09_alarmdb".signal.alarmt12;   // falling edge
   "09_alarmdb".signal.alarmt12 := "06_DB_MOTORS".Rab.Nas29_5;
   IF #_w1 THEN "09_alarmdb".signal_hmi := 12; END_IF;
END_REGION

REGION Network 13
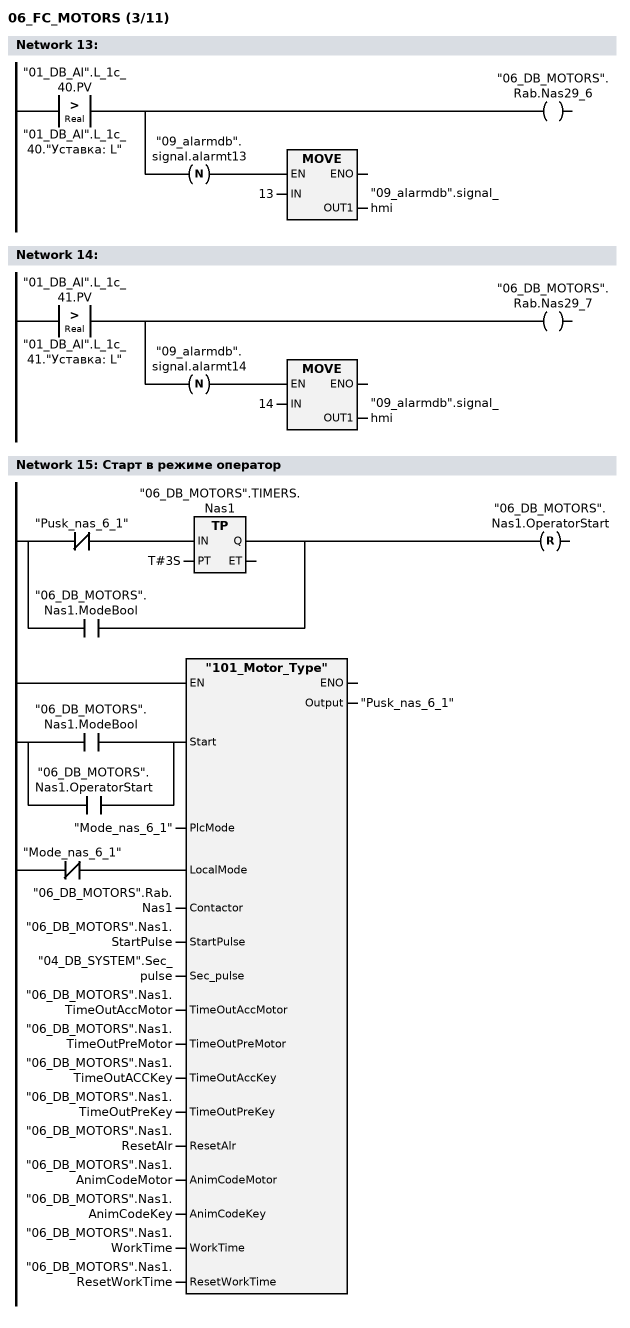
   RUNG wire#powerrail
      { S7_Templates := "SrcType := Real" } GT_Contact(in1 := "01_DB_AI".L_1c_40.PV, in2 := "01_DB_AI".L_1c_40."Уставка: L")
      wire#w1
      Coil( "06_DB_MOTORS".Rab.Nas29_6 )
   END_RUNG
   RUNG wire#w1
      N_Trig( "09_alarmdb".signal.alarmt13 )
      Move(in := 13, out1 => "09_alarmdb".signal_hmi)
   END_RUNG
   // the same network as SCL:
   "06_DB_MOTORS".Rab.Nas29_6 := "01_DB_AI".L_1c_40.PV > "01_DB_AI".L_1c_40."Уставка: L";
   #_w1 := NOT "06_DB_MOTORS".Rab.Nas29_6 AND "09_alarmdb".signal.alarmt13;   // falling edge
   "09_alarmdb".signal.alarmt13 := "06_DB_MOTORS".Rab.Nas29_6;
   IF #_w1 THEN "09_alarmdb".signal_hmi := 13; END_IF;
END_REGION

REGION Network 14
   RUNG wire#powerrail
      { S7_Templates := "SrcType := Real" } GT_Contact(in1 := "01_DB_AI".L_1c_41.PV, in2 := "01_DB_AI".L_1c_41."Уставка: L")
      wire#w1
      Coil( "06_DB_MOTORS".Rab.Nas29_7 )
   END_RUNG
   RUNG wire#w1
      N_Trig( "09_alarmdb".signal.alarmt14 )
      Move(in := 14, out1 => "09_alarmdb".signal_hmi)
   END_RUNG
   // the same network as SCL:
   "06_DB_MOTORS".Rab.Nas29_7 := "01_DB_AI".L_1c_41.PV > "01_DB_AI".L_1c_41."Уставка: L";
   #_w1 := NOT "06_DB_MOTORS".Rab.Nas29_7 AND "09_alarmdb".signal.alarmt14;   // falling edge
   "09_alarmdb".signal.alarmt14 := "06_DB_MOTORS".Rab.Nas29_7;
   IF #_w1 THEN "09_alarmdb".signal_hmi := 14; END_IF;
END_REGION

REGION Network 15: Старт в режиме оператор
   "06_DB_MOTORS".TIMERS.Nas1.TP(IN := NOT "Pusk_nas_6_1", PT := T#3S);
   IF "06_DB_MOTORS".TIMERS.Nas1.Q OR "06_DB_MOTORS".Nas1.ModeBool THEN
       "06_DB_MOTORS".Nas1.OperatorStart := FALSE;
   END_IF;
   "101_Motor_Type"(Start := "06_DB_MOTORS".Nas1.ModeBool OR "06_DB_MOTORS".Nas1.OperatorStart,
                    PlcMode := "Mode_nas_6_1",
                    LocalMode := NOT "Mode_nas_6_1",
                    Contactor := "06_DB_MOTORS".Rab.Nas1,
                    StartPulse := "06_DB_MOTORS".Nas1.StartPulse,
                    Sec_pulse := "04_DB_SYSTEM".Sec_pulse,
                    TimeOutAccMotor := "06_DB_MOTORS".Nas1.TimeOutAccMotor,
                    TimeOutPreMotor := "06_DB_MOTORS".Nas1.TimeOutPreMotor,
                    TimeOutAccKey := "06_DB_MOTORS".Nas1.TimeOutACCKey,
                    TimeOutPreKey := "06_DB_MOTORS".Nas1.TimeOutPreKey,
                    ResetAlr := "06_DB_MOTORS".Nas1.ResetAlr,
                    AnimCodeMotor := "06_DB_MOTORS".Nas1.AnimCodeMotor,
                    AnimCodeKey := "06_DB_MOTORS".Nas1.AnimCodeKey,
                    WorkTime := "06_DB_MOTORS".Nas1.WorkTime,
                    ResetWorkTime := "06_DB_MOTORS".Nas1.ResetWorkTime,
                    Output => "Pusk_nas_6_1");
END_REGION

REGION Network 16: Старт в режиме оператор